(* Logix 5000 project; controller FV vendor 1 type 14 code 217 rev 31.11; software revision 31.00; part 6 of 63 *)
(* tags used below, declared in another part *)
   Alarm_Reset : BOOL;
   Analog_Fault_No : DINT;
   Analog_Simulation_Enabled : BOOL;
   Default_Check_Time : DINT;
   FR_FV26_LTX01_AI : PlantItem;   // FV26_LTX01
   FR_FV26_LTX01_AI_RawInput : ALIAS FOR RIO_Rack_2:2:I.Ch01Data;   // Real Analog Input , Do Not Use In Code
   FR_FV26_PTX01_AI : PlantItem;   // FV26_PTX01
   FR_FV26_PTX01_AI_RawInput : ALIAS FOR RIO_Rack_2:2:I.Ch00Data;   // Real Analog Input , Do Not Use In Code
   FR_FV27_LTX01_AI : PlantItem;   // FV27_LTX01
   FR_FV27_LTX01_AI_RawInput : ALIAS FOR RIO_Rack_2:2:I.Ch03Data;   // Real Analog Input , Do Not Use In Code
   FR_FV27_PTX01_AI : PlantItem;   // FV27_PTX01
   FR_FV27_PTX01_AI_RawInput : ALIAS FOR RIO_Rack_2:2:I.Ch02Data;   // Real Analog Input , Do Not Use In Code
   FR_FV28_LTX01_AI : PlantItem;   // FV28_LTX01
   FR_FV28_LTX01_AI_RawInput : ALIAS FOR RIO_Rack_2:2:I.Ch05Data;   // Real Analog Input , Do Not Use In Code
   FR_FV28_PTX01_AI : PlantItem;   // FV28_PTX01
   FR_FV28_PTX01_AI_RawInput : ALIAS FOR RIO_Rack_2:2:I.Ch04Data;   // Real Analog Input , Do Not Use In Code
   FR_FV29_LTX01_AI : PlantItem;   // FV29_LTX01
   FR_FV29_LTX01_AI_RawInput : ALIAS FOR RIO_Rack_2:2:I.Ch07Data;   // Real Analog Input , Do Not Use In Code
   FR_FV29_PTX01_AI : PlantItem;   // FV29_PTX01
   FR_FV29_PTX01_AI_RawInput : ALIAS FOR RIO_Rack_2:2:I.Ch06Data;   // Real Analog Input , Do Not Use In Code
   FR_FV30_LTX01_AI : PlantItem;   // FV30_LTX01
   FR_FV30_LTX01_AI_RawInput : ALIAS FOR RIO_Rack_2:2:I.Ch09Data;   // Real Analog Input , Do Not Use In Code
   FR_FV30_PTX01_AI : PlantItem;   // FV30_PTX01
   FR_FV30_PTX01_AI_RawInput : ALIAS FOR RIO_Rack_2:2:I.Ch08Data;   // Real Analog Input , Do Not Use In Code
   FR_FV31_LTX01_AI : PlantItem;   // FV31_LTX01
   FR_FV31_LTX01_AI_RawInput : ALIAS FOR RIO_Rack_2:2:I.Ch11Data;   // Real Analog Input , Do Not Use In Code
   FR_FV31_PTX01_AI : PlantItem;   // FV31_PTX01
   FR_FV31_PTX01_AI_RawInput : ALIAS FOR RIO_Rack_2:2:I.Ch10Data;   // Real Analog Input , Do Not Use In Code
   FR_N200 : INT[265];   // ANALOG_IN Analog Inputs
   FR_N210 : INT[265];   // ANALOG_OUT Analog Outputs
   FR_N99 : INT[265];   // COMMENT Comment Lines
   FR_YM_P01_AO : PlantItem;   // YM_P01
   FR_YM_P01_AO_RawOutput : ALIAS FOR RIO_Rack_2:1:O.Ch0Data;   // Real Analog Input , Do Not Use In Code
   FR_YM_P02_AO : PlantItem;   // YM_P02
   FR_YM_P02_AO_RawOutput : ALIAS FOR RIO_Rack_2:1:O.Ch1Data;   // Real Analog Input , Do Not Use In Code
   FR_YM_P03_AO : PlantItem;   // YM_P03
   FR_YM_P03_AO_RawOutput : ALIAS FOR RIO_Rack_2:1:O.Ch2Data;   // Real Analog Input , Do Not Use In Code
   One_Second_One_Scan : ALIAS FOR One_Second_1_scan;
   overrange_RIO_analog_value : REAL;
   underrange_RIO_analog_value : REAL;
(* FR_Common, continued *)

ROUTINE FR_ANALOGI_200   (* ladder *)
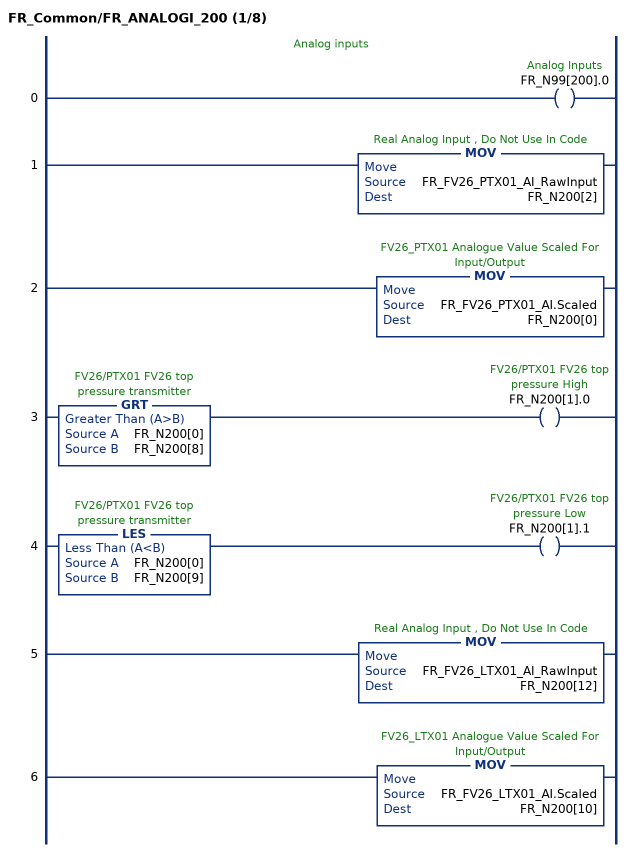
   // Analog inputs
   0: OTE(FR_N99[200].0);
   1: MOV(FR_FV26_PTX01_AI_RawInput,FR_N200[2]);
   2: MOV(FR_FV26_PTX01_AI.Scaled,FR_N200[0]);
   3: GRT(FR_N200[0],FR_N200[8])OTE(FR_N200[1].0);
   4: LES(FR_N200[0],FR_N200[9])OTE(FR_N200[1].1);
   5: MOV(FR_FV26_LTX01_AI_RawInput,FR_N200[12]);
   6: MOV(FR_FV26_LTX01_AI.Scaled,FR_N200[10]);
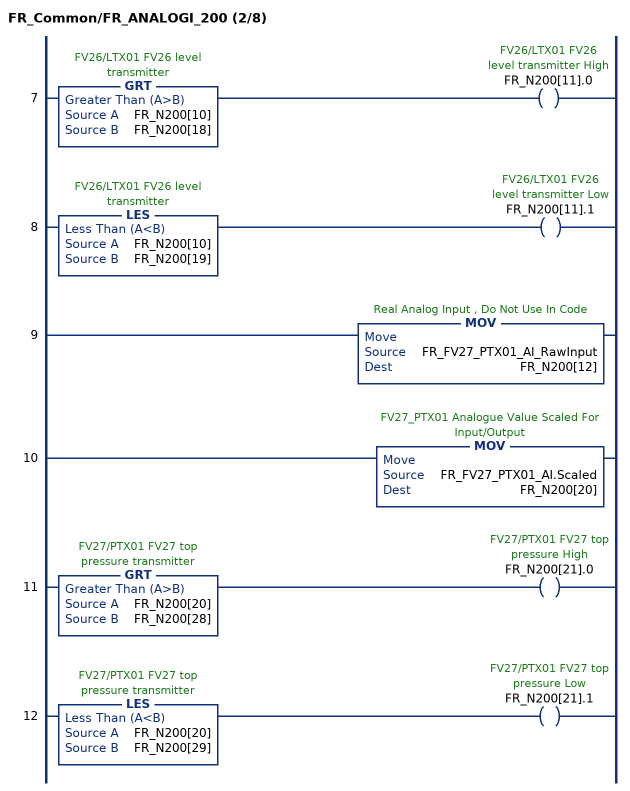
   7: GRT(FR_N200[10],FR_N200[18])OTE(FR_N200[11].0);
   8: LES(FR_N200[10],FR_N200[19])OTE(FR_N200[11].1);
   9: MOV(FR_FV27_PTX01_AI_RawInput,FR_N200[12]);
   10: MOV(FR_FV27_PTX01_AI.Scaled,FR_N200[20]);
   11: GRT(FR_N200[20],FR_N200[28])OTE(FR_N200[21].0);
   12: LES(FR_N200[20],FR_N200[29])OTE(FR_N200[21].1);
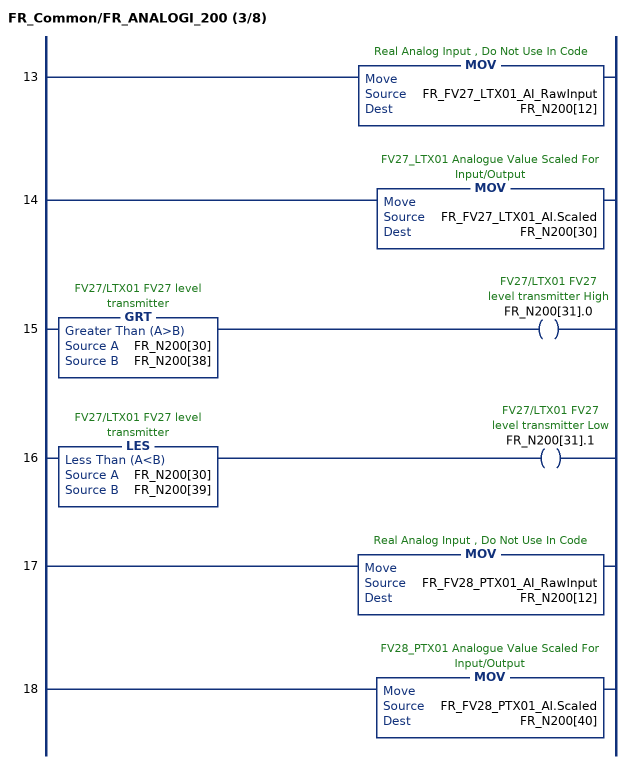
   13: MOV(FR_FV27_LTX01_AI_RawInput,FR_N200[12]);
   14: MOV(FR_FV27_LTX01_AI.Scaled,FR_N200[30]);
   15: GRT(FR_N200[30],FR_N200[38])OTE(FR_N200[31].0);
   16: LES(FR_N200[30],FR_N200[39])OTE(FR_N200[31].1);
   17: MOV(FR_FV28_PTX01_AI_RawInput,FR_N200[12]);
   18: MOV(FR_FV28_PTX01_AI.Scaled,FR_N200[40]);
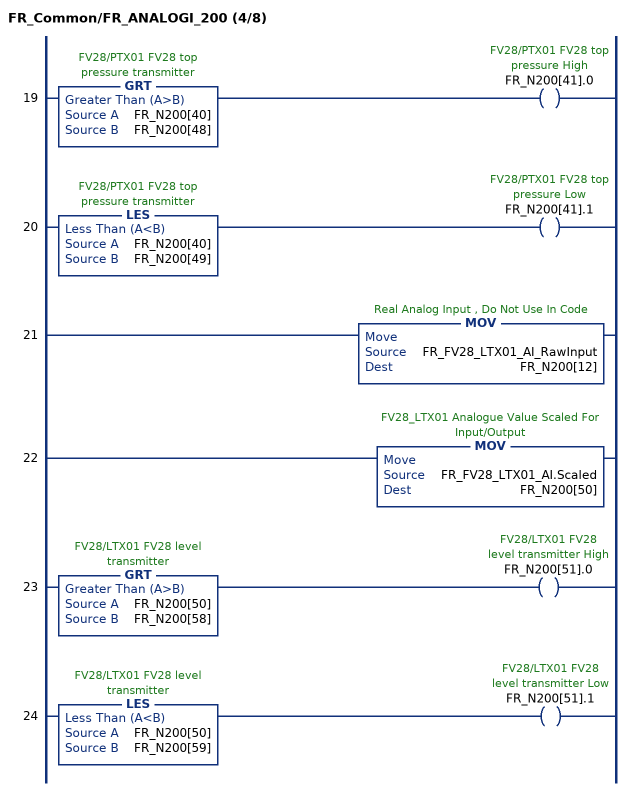
   19: GRT(FR_N200[40],FR_N200[48])OTE(FR_N200[41].0);
   20: LES(FR_N200[40],FR_N200[49])OTE(FR_N200[41].1);
   21: MOV(FR_FV28_LTX01_AI_RawInput,FR_N200[12]);
   22: MOV(FR_FV28_LTX01_AI.Scaled,FR_N200[50]);
   23: GRT(FR_N200[50],FR_N200[58])OTE(FR_N200[51].0);
   24: LES(FR_N200[50],FR_N200[59])OTE(FR_N200[51].1);
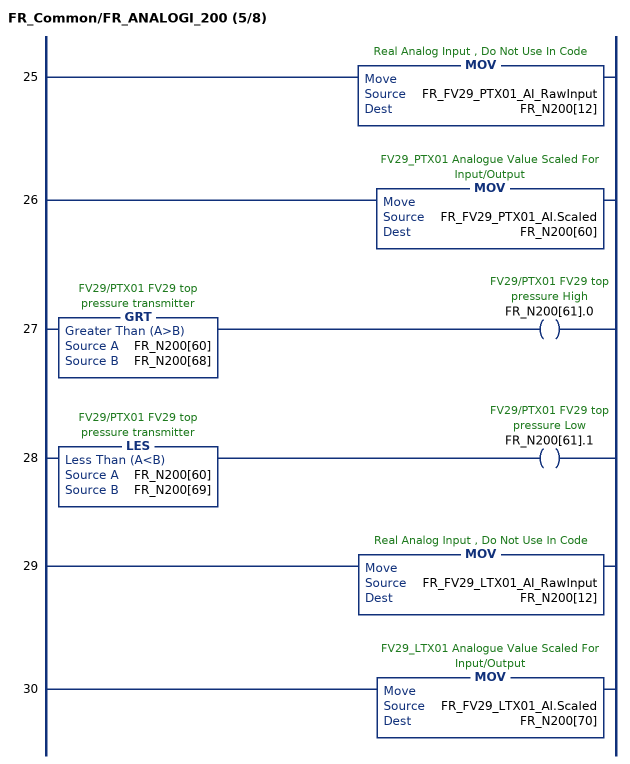
   25: MOV(FR_FV29_PTX01_AI_RawInput,FR_N200[12]);
   26: MOV(FR_FV29_PTX01_AI.Scaled,FR_N200[60]);
   27: GRT(FR_N200[60],FR_N200[68])OTE(FR_N200[61].0);
   28: LES(FR_N200[60],FR_N200[69])OTE(FR_N200[61].1);
   29: MOV(FR_FV29_LTX01_AI_RawInput,FR_N200[12]);
   30: MOV(FR_FV29_LTX01_AI.Scaled,FR_N200[70]);
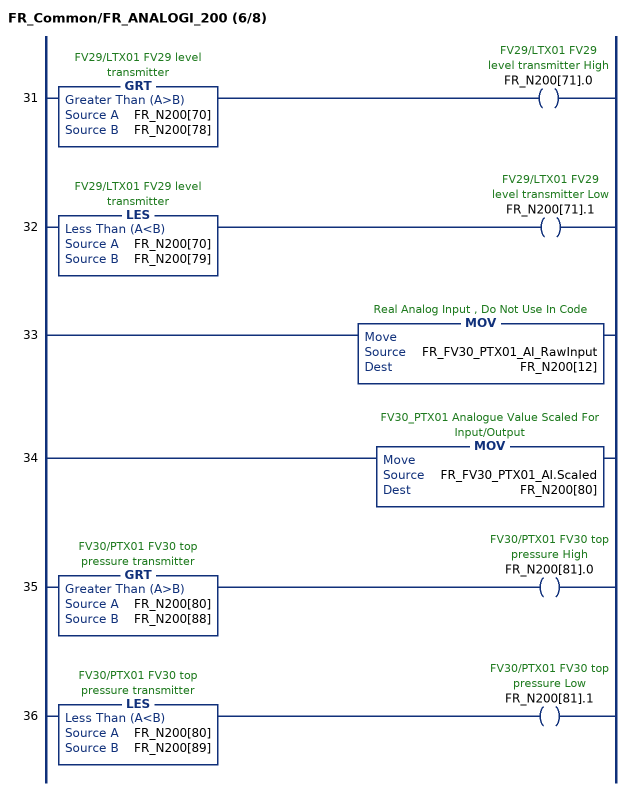
   31: GRT(FR_N200[70],FR_N200[78])OTE(FR_N200[71].0);
   32: LES(FR_N200[70],FR_N200[79])OTE(FR_N200[71].1);
   33: MOV(FR_FV30_PTX01_AI_RawInput,FR_N200[12]);
   34: MOV(FR_FV30_PTX01_AI.Scaled,FR_N200[80]);
   35: GRT(FR_N200[80],FR_N200[88])OTE(FR_N200[81].0);
   36: LES(FR_N200[80],FR_N200[89])OTE(FR_N200[81].1);
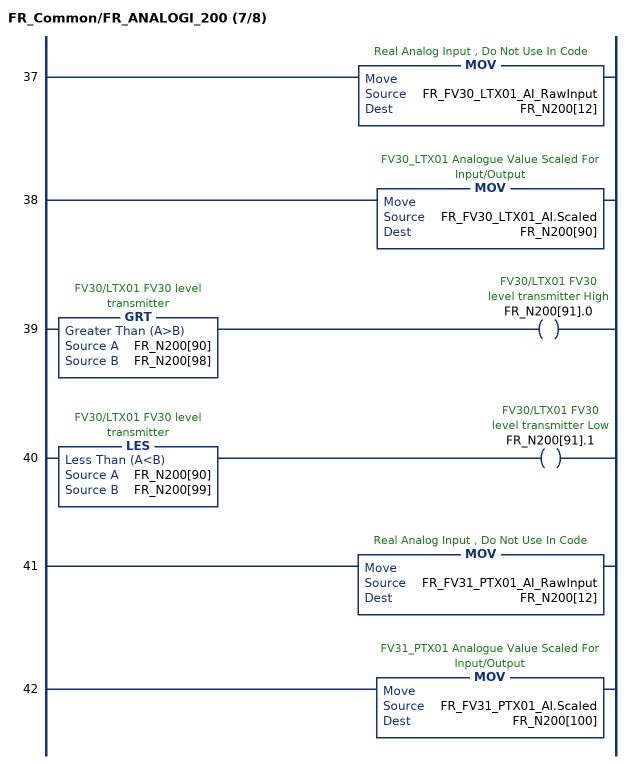
   37: MOV(FR_FV30_LTX01_AI_RawInput,FR_N200[12]);
   38: MOV(FR_FV30_LTX01_AI.Scaled,FR_N200[90]);
   39: GRT(FR_N200[90],FR_N200[98])OTE(FR_N200[91].0);
   40: LES(FR_N200[90],FR_N200[99])OTE(FR_N200[91].1);
   41: MOV(FR_FV31_PTX01_AI_RawInput,FR_N200[12]);
   42: MOV(FR_FV31_PTX01_AI.Scaled,FR_N200[100]);
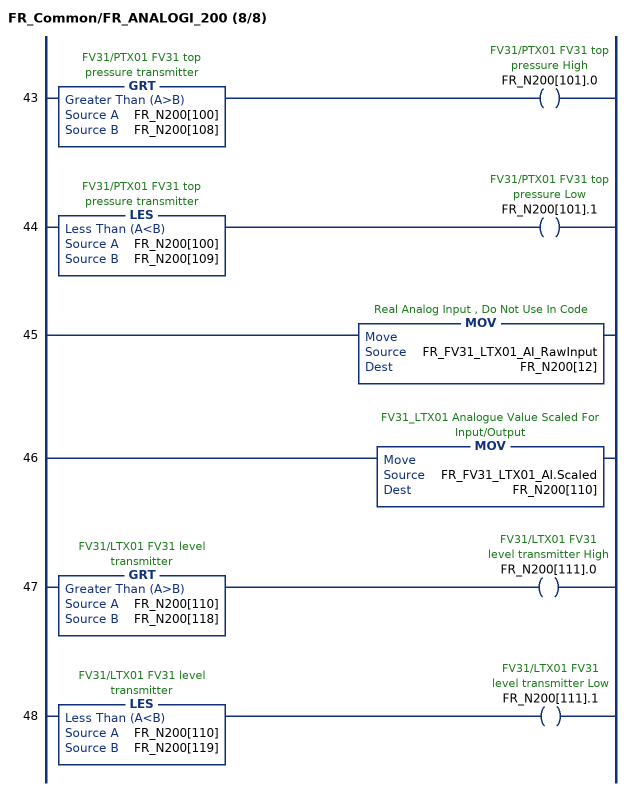
   43: GRT(FR_N200[100],FR_N200[108])OTE(FR_N200[101].0);
   44: LES(FR_N200[100],FR_N200[109])OTE(FR_N200[101].1);
   45: MOV(FR_FV31_LTX01_AI_RawInput,FR_N200[12]);
   46: MOV(FR_FV31_LTX01_AI.Scaled,FR_N200[110]);
   47: GRT(FR_N200[110],FR_N200[118])OTE(FR_N200[111].0);
   48: LES(FR_N200[110],FR_N200[119])OTE(FR_N200[111].1);
END_ROUTINE

ROUTINE FR_ANALOGO_210   (* ladder *)
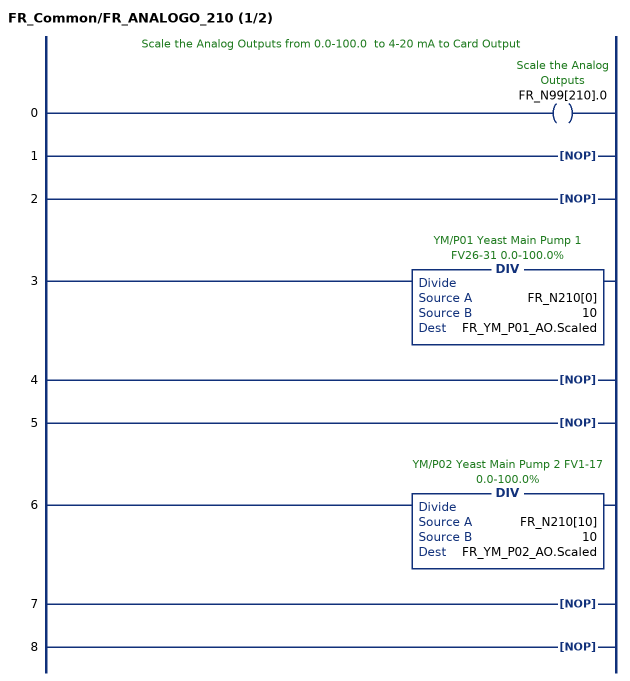
   // Scale the Analog Outputs from 0.0-100.0  to 4-20 mA to Card Output
   0: OTE(FR_N99[210].0);
   1: NOP();
   2: NOP();
   3: DIV(FR_N210[0],10,FR_YM_P01_AO.Scaled);
   4: NOP();
   5: NOP();
   6: DIV(FR_N210[10],10,FR_YM_P02_AO.Scaled);
   7: NOP();
   8: NOP();
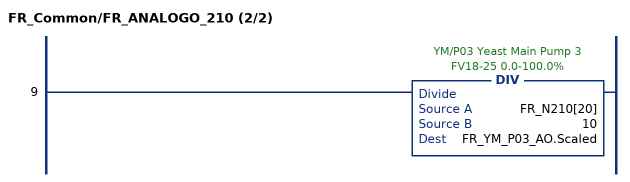
   9: DIV(FR_N210[20],10,FR_YM_P03_AO.Scaled);
END_ROUTINE

ROUTINE FR_Analogs   (* ladder *)
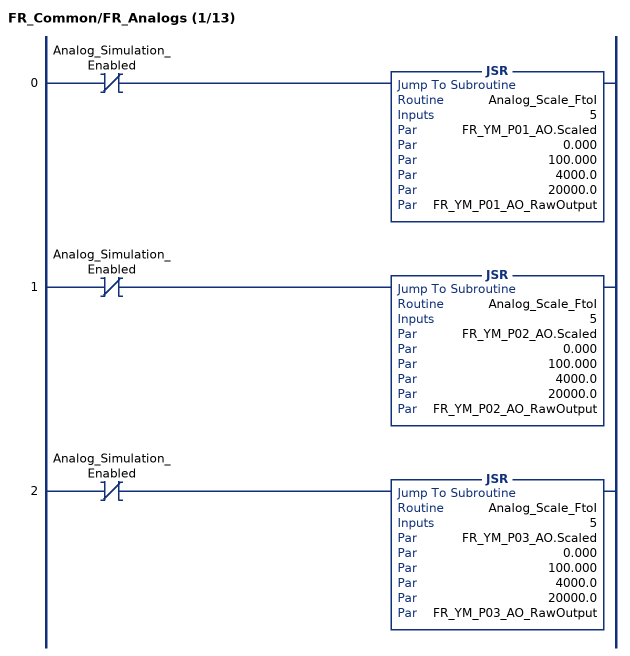
   0: XIO(Analog_Simulation_Enabled)JSR(Analog_Scale_FtoI,5,FR_YM_P01_AO.Scaled,0.000,100.000,4000.0,20000.0,FR_YM_P01_AO_RawOutput);
   1: XIO(Analog_Simulation_Enabled)JSR(Analog_Scale_FtoI,5,FR_YM_P02_AO.Scaled,0.000,100.000,4000.0,20000.0,FR_YM_P02_AO_RawOutput);
   2: XIO(Analog_Simulation_Enabled)JSR(Analog_Scale_FtoI,5,FR_YM_P03_AO.Scaled,0.000,100.000,4000.0,20000.0,FR_YM_P03_AO_RawOutput);
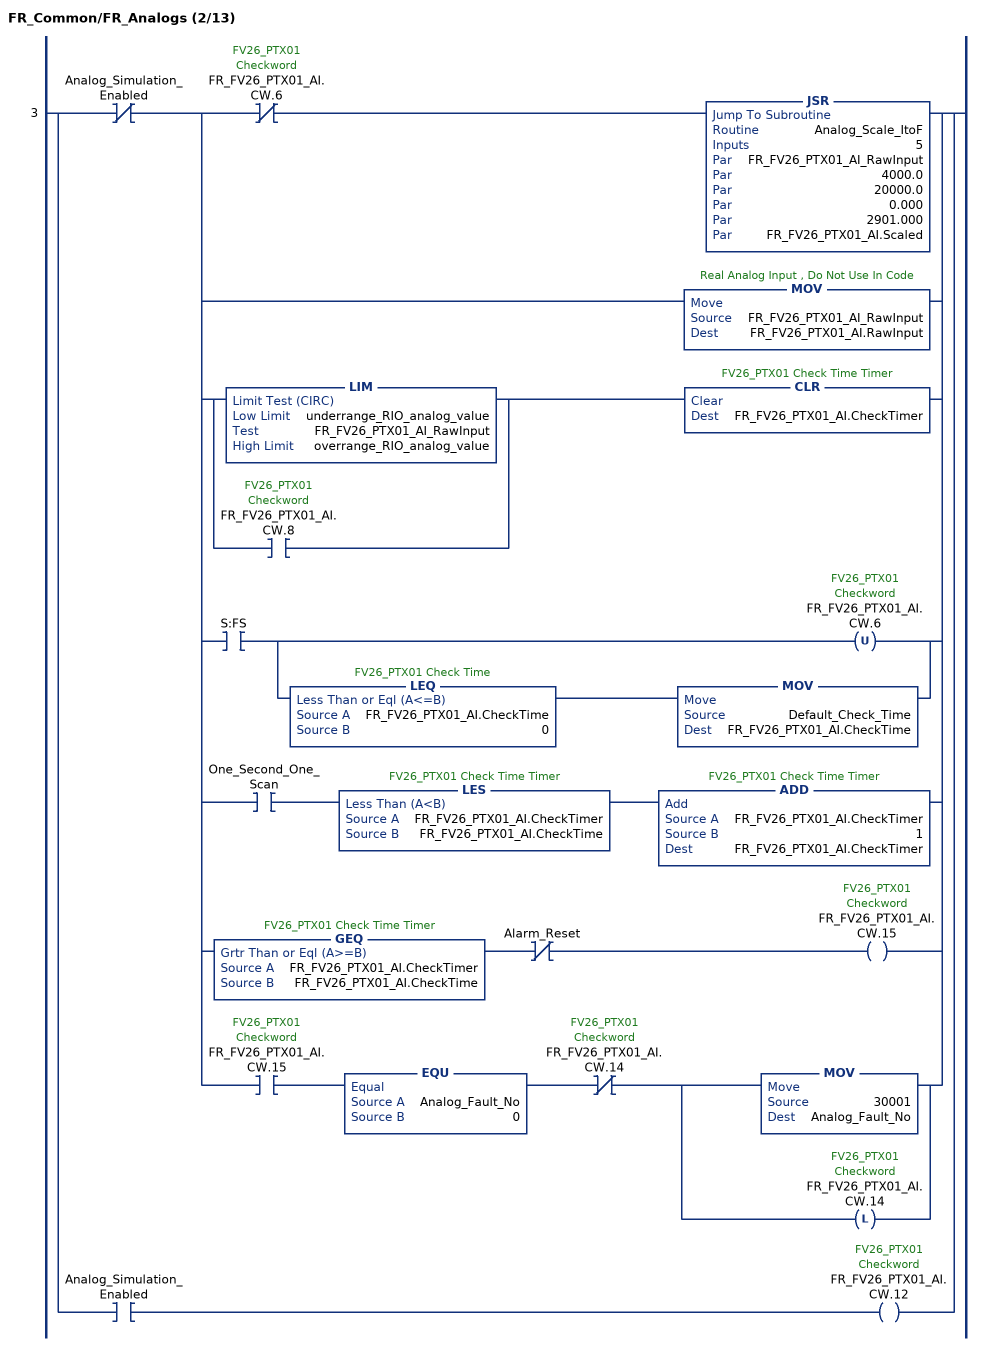
   3: [XIO(Analog_Simulation_Enabled) [XIO(FR_FV26_PTX01_AI.CW.6) JSR(Analog_Scale_ItoF,5,FR_FV26_PTX01_AI_RawInput,4000.0,20000.0,0.000,2901.000,FR_FV26_PTX01_AI.Scaled) ,MOV(FR_FV26_PTX01_AI_RawInput,FR_FV26_PTX01_AI.RawInput) ,[LIM(underrange_RIO_analog_value,FR_FV26_PTX01_AI_RawInput,overrange_RIO_analog_value) ,XIC(FR_FV26_PTX01_AI.CW.8) ] CLR(FR_FV26_PTX01_AI.CheckTimer) ,XIC(S:FS) [OTU(FR_FV26_PTX01_AI.CW.6) ,LEQ(FR_FV26_PTX01_AI.CheckTime,0) MOV(Default_Check_Time,FR_FV26_PTX01_AI.CheckTime) ] ,XIC(One_Second_One_Scan) LES(FR_FV26_PTX01_AI.CheckTimer,FR_FV26_PTX01_AI.CheckTime) ADD(FR_FV26_PTX01_AI.CheckTimer,1,FR_FV26_PTX01_AI.CheckTimer) ,GEQ(FR_FV26_PTX01_AI.CheckTimer,FR_FV26_PTX01_AI.CheckTime) XIO(Alarm_Reset) OTE(FR_FV26_PTX01_AI.CW.15) ,XIC(FR_FV26_PTX01_AI.CW.15) EQU(Analog_Fault_No,0) XIO(FR_FV26_PTX01_AI.CW.14) [MOV(30001,Analog_Fault_No) ,OTL(FR_FV26_PTX01_AI.CW.14) ] ] ,XIC(Analog_Simulation_Enabled) OTE(FR_FV26_PTX01_AI.CW.12) ];
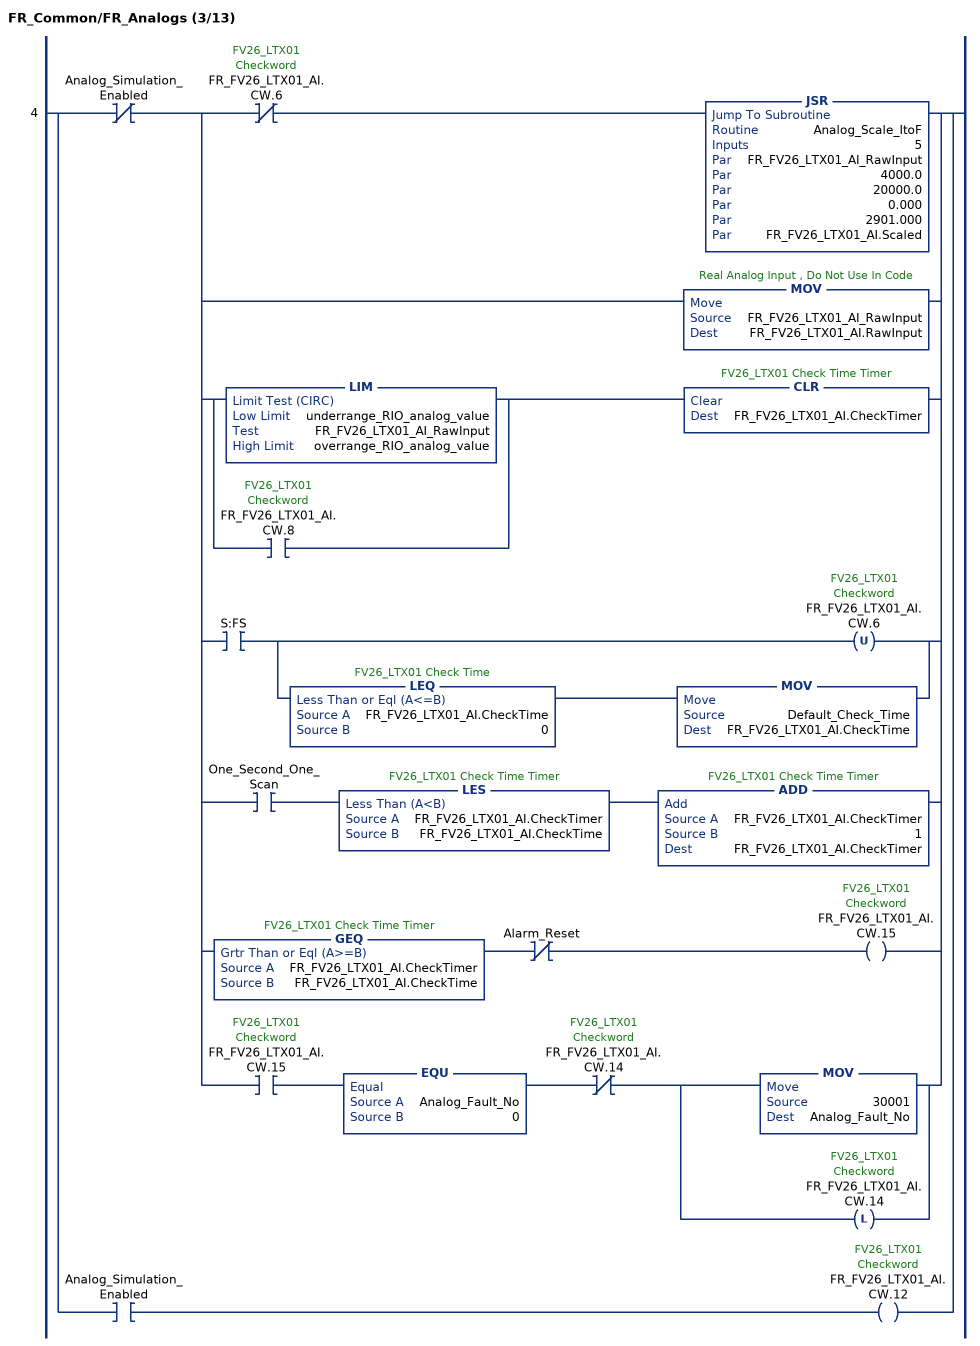
   4: [XIO(Analog_Simulation_Enabled) [XIO(FR_FV26_LTX01_AI.CW.6) JSR(Analog_Scale_ItoF,5,FR_FV26_LTX01_AI_RawInput,4000.0,20000.0,0.000,2901.000,FR_FV26_LTX01_AI.Scaled) ,MOV(FR_FV26_LTX01_AI_RawInput,FR_FV26_LTX01_AI.RawInput) ,[LIM(underrange_RIO_analog_value,FR_FV26_LTX01_AI_RawInput,overrange_RIO_analog_value) ,XIC(FR_FV26_LTX01_AI.CW.8) ] CLR(FR_FV26_LTX01_AI.CheckTimer) ,XIC(S:FS) [OTU(FR_FV26_LTX01_AI.CW.6) ,LEQ(FR_FV26_LTX01_AI.CheckTime,0) MOV(Default_Check_Time,FR_FV26_LTX01_AI.CheckTime) ] ,XIC(One_Second_One_Scan) LES(FR_FV26_LTX01_AI.CheckTimer,FR_FV26_LTX01_AI.CheckTime) ADD(FR_FV26_LTX01_AI.CheckTimer,1,FR_FV26_LTX01_AI.CheckTimer) ,GEQ(FR_FV26_LTX01_AI.CheckTimer,FR_FV26_LTX01_AI.CheckTime) XIO(Alarm_Reset) OTE(FR_FV26_LTX01_AI.CW.15) ,XIC(FR_FV26_LTX01_AI.CW.15) EQU(Analog_Fault_No,0) XIO(FR_FV26_LTX01_AI.CW.14) [MOV(30001,Analog_Fault_No) ,OTL(FR_FV26_LTX01_AI.CW.14) ] ] ,XIC(Analog_Simulation_Enabled) OTE(FR_FV26_LTX01_AI.CW.12) ];
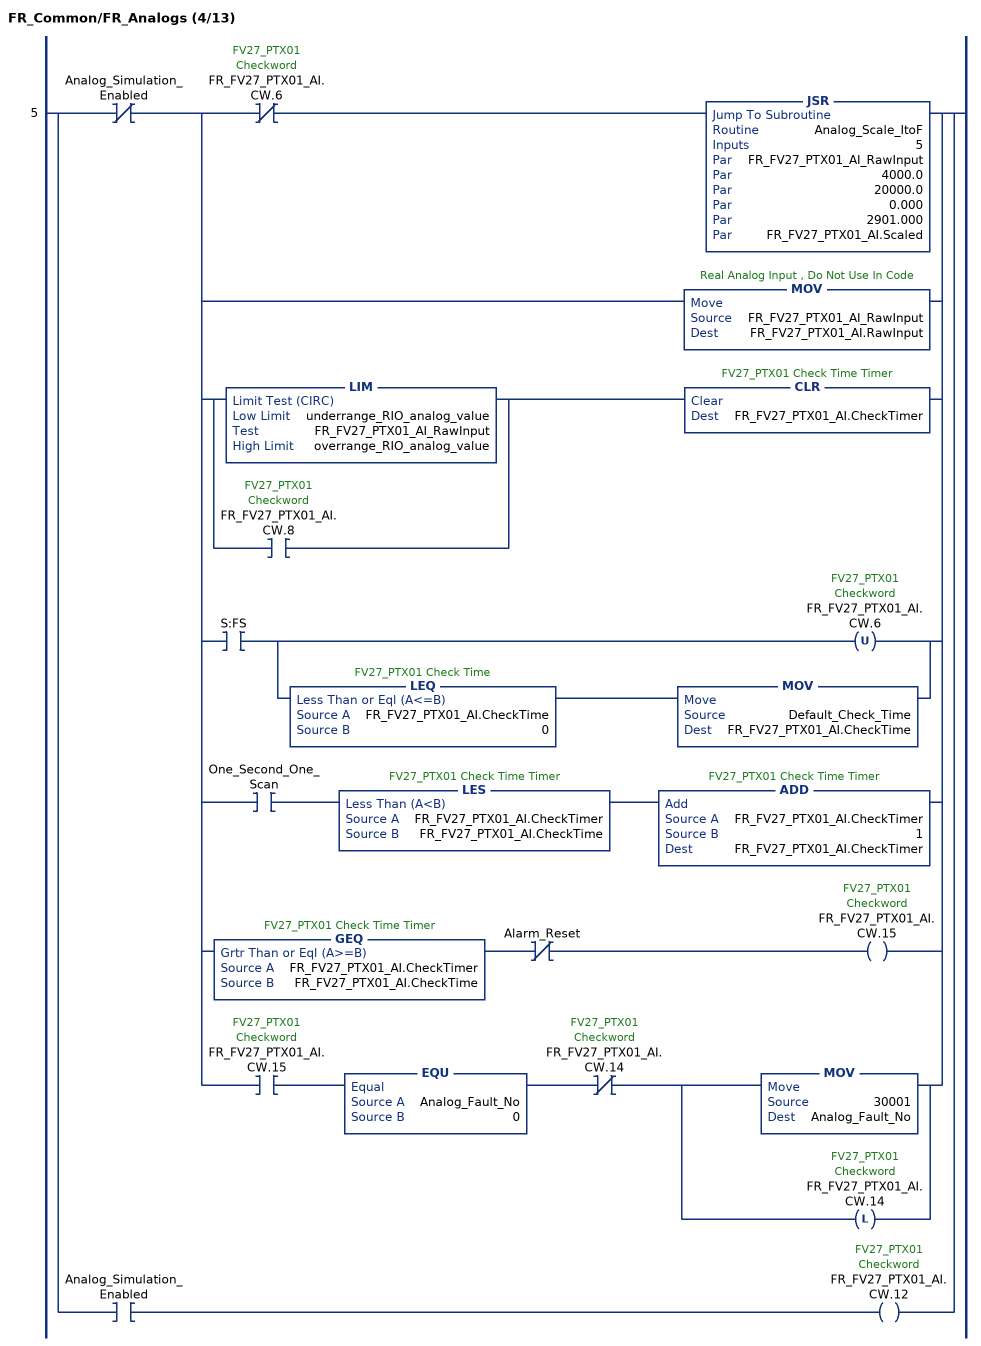
   5: [XIO(Analog_Simulation_Enabled) [XIO(FR_FV27_PTX01_AI.CW.6) JSR(Analog_Scale_ItoF,5,FR_FV27_PTX01_AI_RawInput,4000.0,20000.0,0.000,2901.000,FR_FV27_PTX01_AI.Scaled) ,MOV(FR_FV27_PTX01_AI_RawInput,FR_FV27_PTX01_AI.RawInput) ,[LIM(underrange_RIO_analog_value,FR_FV27_PTX01_AI_RawInput,overrange_RIO_analog_value) ,XIC(FR_FV27_PTX01_AI.CW.8) ] CLR(FR_FV27_PTX01_AI.CheckTimer) ,XIC(S:FS) [OTU(FR_FV27_PTX01_AI.CW.6) ,LEQ(FR_FV27_PTX01_AI.CheckTime,0) MOV(Default_Check_Time,FR_FV27_PTX01_AI.CheckTime) ] ,XIC(One_Second_One_Scan) LES(FR_FV27_PTX01_AI.CheckTimer,FR_FV27_PTX01_AI.CheckTime) ADD(FR_FV27_PTX01_AI.CheckTimer,1,FR_FV27_PTX01_AI.CheckTimer) ,GEQ(FR_FV27_PTX01_AI.CheckTimer,FR_FV27_PTX01_AI.CheckTime) XIO(Alarm_Reset) OTE(FR_FV27_PTX01_AI.CW.15) ,XIC(FR_FV27_PTX01_AI.CW.15) EQU(Analog_Fault_No,0) XIO(FR_FV27_PTX01_AI.CW.14) [MOV(30001,Analog_Fault_No) ,OTL(FR_FV27_PTX01_AI.CW.14) ] ] ,XIC(Analog_Simulation_Enabled) OTE(FR_FV27_PTX01_AI.CW.12) ];